(* Logix 5000 project; controller UOWHF_Vary Emulate 5570 rev 30.12; software revision 30.00; part 13 of 13 *)
(* tags used below, declared in another part *)
   UOWHF_Add_c : DINT;
   UOWHF_i : DINT;
   UOWHF_InputLen : DINT;
   UOWHF_InputMaxInd : DINT;
   UOWHF_Msg : DINT[16];
   UOWHF_OutputMaxInd : DINT;
   UOWHF_Result : DINT[17];
   UOWHF_Vary_BlkNum : DINT;
   UOWHF_Vary_i : DINT;
   UOWHF_Vary_j : DINT;
   UOWHF_Vary_Message : DINT[512];
   UOWHF_Vary_MsgLen : DINT;
   UOWHF_Vary_z : DINT;
   UOWHF_VaryLen : DINT;
   UOWHF_Ver : DINT;
(* MainProgram, continued *)

   		UOWHF_Add_c.7:=UOWHF_Result[7].31;
   		UOWHF_Result[7].31:=0;
   		UOWHF_Result[8]:=UOWHF_Result[8] + 1529564597+UOWHF_Add_c;
   		UOWHF_Add_c.8:=UOWHF_Result[8].31;
   		UOWHF_Result[8].31:=0;
   	End_If;
   	If UOWHF_Msg[15].[5] Then
   		UOWHF_Result[0]:=UOWHF_Result[0] + 534622081+UOWHF_Add_c;
   		UOWHF_Add_c.0:=UOWHF_Result[0].31;
   		UOWHF_Result[0].31:=0;
   		UOWHF_Result[1]:=UOWHF_Result[1] + 1054997605+UOWHF_Add_c;
   		UOWHF_Add_c.1:=UOWHF_Result[1].31;
   		UOWHF_Result[1].31:=0;
   		UOWHF_Result[2]:=UOWHF_Result[2] + 944898288+UOWHF_Add_c;
   		UOWHF_Add_c.2:=UOWHF_Result[2].31;
   		UOWHF_Result[2].31:=0;
   		UOWHF_Result[3]:=UOWHF_Result[3] + 811676453+UOWHF_Add_c;
   		UOWHF_Add_c.3:=UOWHF_Result[3].31;
   		UOWHF_Result[3].31:=0;
   		UOWHF_Result[4]:=UOWHF_Result[4] + 1761848356+UOWHF_Add_c;
   		UOWHF_Add_c.4:=UOWHF_Result[4].31;
   		UOWHF_Result[4].31:=0;
   		UOWHF_Result[5]:=UOWHF_Result[5] + 163403387+UOWHF_Add_c;
   		UOWHF_Add_c.5:=UOWHF_Result[5].31;
   		UOWHF_Result[5].31:=0;
   		UOWHF_Result[6]:=UOWHF_Result[6] + 606196183+UOWHF_Add_c;
   		UOWHF_Add_c.6:=UOWHF_Result[6].31;
   		UOWHF_Result[6].31:=0;
   		UOWHF_Result[7]:=UOWHF_Result[7] + 2030634477+UOWHF_Add_c;
   		UOWHF_Add_c.7:=UOWHF_Result[7].31;
   		UOWHF_Result[7].31:=0;
   		UOWHF_Result[8]:=UOWHF_Result[8] + 457492181+UOWHF_Add_c;
   		UOWHF_Add_c.8:=UOWHF_Result[8].31;
   		UOWHF_Result[8].31:=0;
   	End_If;
   	If UOWHF_Msg[15].[6] Then
   		UOWHF_Result[0]:=UOWHF_Result[0] + 1563595876+UOWHF_Add_c;
   		UOWHF_Add_c.0:=UOWHF_Result[0].31;
   		UOWHF_Result[0].31:=0;
   		UOWHF_Result[1]:=UOWHF_Result[1] + 921060794+UOWHF_Add_c;
   		UOWHF_Add_c.1:=UOWHF_Result[1].31;
   		UOWHF_Result[1].31:=0;
   		UOWHF_Result[2]:=UOWHF_Result[2] + 1052970481+UOWHF_Add_c;
   		UOWHF_Add_c.2:=UOWHF_Result[2].31;
   		UOWHF_Result[2].31:=0;
   		UOWHF_Result[3]:=UOWHF_Result[3] + 657088809+UOWHF_Add_c;
   		UOWHF_Add_c.3:=UOWHF_Result[3].31;
   		UOWHF_Result[3].31:=0;
   		UOWHF_Result[4]:=UOWHF_Result[4] + 107170927+UOWHF_Add_c;
   		UOWHF_Add_c.4:=UOWHF_Result[4].31;
   		UOWHF_Result[4].31:=0;
   		UOWHF_Result[5]:=UOWHF_Result[5] + 1430973014+UOWHF_Add_c;
   		UOWHF_Add_c.5:=UOWHF_Result[5].31;
   		UOWHF_Result[5].31:=0;
   		UOWHF_Result[6]:=UOWHF_Result[6] + 454401316+UOWHF_Add_c;
   		UOWHF_Add_c.6:=UOWHF_Result[6].31;
   		UOWHF_Result[6].31:=0;
   		UOWHF_Result[7]:=UOWHF_Result[7] + 395129130+UOWHF_Add_c;
   		UOWHF_Add_c.7:=UOWHF_Result[7].31;
   		UOWHF_Result[7].31:=0;
   		UOWHF_Result[8]:=UOWHF_Result[8] + 1072078032+UOWHF_Add_c;
   		UOWHF_Add_c.8:=UOWHF_Result[8].31;
   		UOWHF_Result[8].31:=0;
   	End_If;
   	If UOWHF_Msg[15].[7] Then
   		UOWHF_Result[0]:=UOWHF_Result[0] + 1403391658+UOWHF_Add_c;
   		UOWHF_Add_c.0:=UOWHF_Result[0].31;
   		UOWHF_Result[0].31:=0;
   		UOWHF_Result[1]:=UOWHF_Result[1] + 1796223182+UOWHF_Add_c;
   		UOWHF_Add_c.1:=UOWHF_Result[1].31;
   		UOWHF_Result[1].31:=0;
   		UOWHF_Result[2]:=UOWHF_Result[2] + 960792761+UOWHF_Add_c;
   		UOWHF_Add_c.2:=UOWHF_Result[2].31;
   		UOWHF_Result[2].31:=0;
   		UOWHF_Result[3]:=UOWHF_Result[3] + 288040454+UOWHF_Add_c;
   		UOWHF_Add_c.3:=UOWHF_Result[3].31;
   		UOWHF_Result[3].31:=0;
   		UOWHF_Result[4]:=UOWHF_Result[4] + 356603480+UOWHF_Add_c;
   		UOWHF_Add_c.4:=UOWHF_Result[4].31;
   		UOWHF_Result[4].31:=0;
   		UOWHF_Result[5]:=UOWHF_Result[5] + 1694776766+UOWHF_Add_c;
   		UOWHF_Add_c.5:=UOWHF_Result[5].31;
   		UOWHF_Result[5].31:=0;
   		UOWHF_Result[6]:=UOWHF_Result[6] + 1001613380+UOWHF_Add_c;
   		UOWHF_Add_c.6:=UOWHF_Result[6].31;
   		UOWHF_Result[6].31:=0;
   		UOWHF_Result[7]:=UOWHF_Result[7] + 1296327921+UOWHF_Add_c;
   		UOWHF_Add_c.7:=UOWHF_Result[7].31;
   		UOWHF_Result[7].31:=0;
   		UOWHF_Result[8]:=UOWHF_Result[8] + 1853983857+UOWHF_Add_c;
   		UOWHF_Add_c.8:=UOWHF_Result[8].31;
   		UOWHF_Result[8].31:=0;
   	End_If;
   	If UOWHF_Msg[15].[8] Then
   		UOWHF_Result[0]:=UOWHF_Result[0] + 1265129415+UOWHF_Add_c;
   		UOWHF_Add_c.0:=UOWHF_Result[0].31;
   		UOWHF_Result[0].31:=0;
   		UOWHF_Result[1]:=UOWHF_Result[1] + 568656446+UOWHF_Add_c;
   		UOWHF_Add_c.1:=UOWHF_Result[1].31;
   		UOWHF_Result[1].31:=0;
   		UOWHF_Result[2]:=UOWHF_Result[2] + 1035914428+UOWHF_Add_c;
   		UOWHF_Add_c.2:=UOWHF_Result[2].31;
   		UOWHF_Result[2].31:=0;
   		UOWHF_Result[3]:=UOWHF_Result[3] + 1838467801+UOWHF_Add_c;
   		UOWHF_Add_c.3:=UOWHF_Result[3].31;
   		UOWHF_Result[3].31:=0;
   		UOWHF_Result[4]:=UOWHF_Result[4] + 852571844+UOWHF_Add_c;
   		UOWHF_Add_c.4:=UOWHF_Result[4].31;
   		UOWHF_Result[4].31:=0;
   		UOWHF_Result[5]:=UOWHF_Result[5] + 811437709+UOWHF_Add_c;
   		UOWHF_Add_c.5:=UOWHF_Result[5].31;
   		UOWHF_Result[5].31:=0;
   		UOWHF_Result[6]:=UOWHF_Result[6] + 2110578431+UOWHF_Add_c;
   		UOWHF_Add_c.6:=UOWHF_Result[6].31;
   		UOWHF_Result[6].31:=0;
   		UOWHF_Result[7]:=UOWHF_Result[7] + 1083369967+UOWHF_Add_c;
   		UOWHF_Add_c.7:=UOWHF_Result[7].31;
   		UOWHF_Result[7].31:=0;
   		UOWHF_Result[8]:=UOWHF_Result[8] + 1040887567+UOWHF_Add_c;
   		UOWHF_Add_c.8:=UOWHF_Result[8].31;
   		UOWHF_Result[8].31:=0;
   	End_If;
   	If UOWHF_Msg[15].[9] Then
   		UOWHF_Result[0]:=UOWHF_Result[0] + 1883016459+UOWHF_Add_c;
   		UOWHF_Add_c.0:=UOWHF_Result[0].31;
   		UOWHF_Result[0].31:=0;
   		UOWHF_Result[1]:=UOWHF_Result[1] + 1109215782+UOWHF_Add_c;
   		UOWHF_Add_c.1:=UOWHF_Result[1].31;
   		UOWHF_Result[1].31:=0;
   		UOWHF_Result[2]:=UOWHF_Result[2] + 692572348+UOWHF_Add_c;
   		UOWHF_Add_c.2:=UOWHF_Result[2].31;
   		UOWHF_Result[2].31:=0;
   		UOWHF_Result[3]:=UOWHF_Result[3] + 357248589+UOWHF_Add_c;
   		UOWHF_Add_c.3:=UOWHF_Result[3].31;
   		UOWHF_Result[3].31:=0;
   		UOWHF_Result[4]:=UOWHF_Result[4] + 495139913+UOWHF_Add_c;
   		UOWHF_Add_c.4:=UOWHF_Result[4].31;
   		UOWHF_Result[4].31:=0;
   		UOWHF_Result[5]:=UOWHF_Result[5] + 1972425862+UOWHF_Add_c;
   		UOWHF_Add_c.5:=UOWHF_Result[5].31;
   		UOWHF_Result[5].31:=0;
   		UOWHF_Result[6]:=UOWHF_Result[6] + 1336574867+UOWHF_Add_c;
   		UOWHF_Add_c.6:=UOWHF_Result[6].31;
   		UOWHF_Result[6].31:=0;
   		UOWHF_Result[7]:=UOWHF_Result[7] + 286906005+UOWHF_Add_c;
   		UOWHF_Add_c.7:=UOWHF_Result[7].31;
   		UOWHF_Result[7].31:=0;
   		UOWHF_Result[8]:=UOWHF_Result[8] + 935997948+UOWHF_Add_c;
   		UOWHF_Add_c.8:=UOWHF_Result[8].31;
   		UOWHF_Result[8].31:=0;
   	End_If;
   	If UOWHF_Msg[15].[10] Then
   		UOWHF_Result[0]:=UOWHF_Result[0] + 406811790+UOWHF_Add_c;
   		UOWHF_Add_c.0:=UOWHF_Result[0].31;
   		UOWHF_Result[0].31:=0;
   		UOWHF_Result[1]:=UOWHF_Result[1] + 1667294919+UOWHF_Add_c;
   		UOWHF_Add_c.1:=UOWHF_Result[1].31;
   		UOWHF_Result[1].31:=0;
   		UOWHF_Result[2]:=UOWHF_Result[2] + 2033524595+UOWHF_Add_c;
   		UOWHF_Add_c.2:=UOWHF_Result[2].31;
   		UOWHF_Result[2].31:=0;
   		UOWHF_Result[3]:=UOWHF_Result[3] + 1349255026+UOWHF_Add_c;
   		UOWHF_Add_c.3:=UOWHF_Result[3].31;
   		UOWHF_Result[3].31:=0;
   		UOWHF_Result[4]:=UOWHF_Result[4] + 10415662+UOWHF_Add_c;
   		UOWHF_Add_c.4:=UOWHF_Result[4].31;
   		UOWHF_Result[4].31:=0;
   		UOWHF_Result[5]:=UOWHF_Result[5] + 2068656448+UOWHF_Add_c;
   		UOWHF_Add_c.5:=UOWHF_Result[5].31;
   		UOWHF_Result[5].31:=0;
   		UOWHF_Result[6]:=UOWHF_Result[6] + 719617830+UOWHF_Add_c;
   		UOWHF_Add_c.6:=UOWHF_Result[6].31;
   		UOWHF_Result[6].31:=0;
   		UOWHF_Result[7]:=UOWHF_Result[7] + 867653174+UOWHF_Add_c;
   		UOWHF_Add_c.7:=UOWHF_Result[7].31;
   		UOWHF_Result[7].31:=0;
   		UOWHF_Result[8]:=UOWHF_Result[8] + 1934472738+UOWHF_Add_c;
   		UOWHF_Add_c.8:=UOWHF_Result[8].31;
   		UOWHF_Result[8].31:=0;
   	End_If;
   	If UOWHF_Msg[15].[11] Then
   		UOWHF_Result[0]:=UOWHF_Result[0] + 165633326+UOWHF_Add_c;
   		UOWHF_Add_c.0:=UOWHF_Result[0].31;
   		UOWHF_Result[0].31:=0;
   		UOWHF_Result[1]:=UOWHF_Result[1] + 53652767+UOWHF_Add_c;
   		UOWHF_Add_c.1:=UOWHF_Result[1].31;
   		UOWHF_Result[1].31:=0;
   		UOWHF_Result[2]:=UOWHF_Result[2] + 1574797324+UOWHF_Add_c;
   		UOWHF_Add_c.2:=UOWHF_Result[2].31;
   		UOWHF_Result[2].31:=0;
   		UOWHF_Result[3]:=UOWHF_Result[3] + 1336775684+UOWHF_Add_c;
   		UOWHF_Add_c.3:=UOWHF_Result[3].31;
   		UOWHF_Result[3].31:=0;
   		UOWHF_Result[4]:=UOWHF_Result[4] + 1894121389+UOWHF_Add_c;
   		UOWHF_Add_c.4:=UOWHF_Result[4].31;
   		UOWHF_Result[4].31:=0;
   		UOWHF_Result[5]:=UOWHF_Result[5] + 1658923569+UOWHF_Add_c;
   		UOWHF_Add_c.5:=UOWHF_Result[5].31;
   		UOWHF_Result[5].31:=0;
   		UOWHF_Result[6]:=UOWHF_Result[6] + 1195345328+UOWHF_Add_c;
   		UOWHF_Add_c.6:=UOWHF_Result[6].31;
   		UOWHF_Result[6].31:=0;
   		UOWHF_Result[7]:=UOWHF_Result[7] + 1912811518+UOWHF_Add_c;
   		UOWHF_Add_c.7:=UOWHF_Result[7].31;
   		UOWHF_Result[7].31:=0;
   		UOWHF_Result[8]:=UOWHF_Result[8] + 826695963+UOWHF_Add_c;
   		UOWHF_Add_c.8:=UOWHF_Result[8].31;
   		UOWHF_Result[8].31:=0;
   	End_If;
   	If UOWHF_Msg[15].[12] Then
   		UOWHF_Result[0]:=UOWHF_Result[0] + 1033530810+UOWHF_Add_c;
   		UOWHF_Add_c.0:=UOWHF_Result[0].31;
   		UOWHF_Result[0].31:=0;
   		UOWHF_Result[1]:=UOWHF_Result[1] + 449682606+UOWHF_Add_c;
   		UOWHF_Add_c.1:=UOWHF_Result[1].31;
   		UOWHF_Result[1].31:=0;
   		UOWHF_Result[2]:=UOWHF_Result[2] + 1100837890+UOWHF_Add_c;
   		UOWHF_Add_c.2:=UOWHF_Result[2].31;
   		UOWHF_Result[2].31:=0;
   		UOWHF_Result[3]:=UOWHF_Result[3] + 721973923+UOWHF_Add_c;
   		UOWHF_Add_c.3:=UOWHF_Result[3].31;
   		UOWHF_Result[3].31:=0;
   		UOWHF_Result[4]:=UOWHF_Result[4] + 2071465357+UOWHF_Add_c;
   		UOWHF_Add_c.4:=UOWHF_Result[4].31;
   		UOWHF_Result[4].31:=0;
   		UOWHF_Result[5]:=UOWHF_Result[5] + 514392075+UOWHF_Add_c;
   		UOWHF_Add_c.5:=UOWHF_Result[5].31;
   		UOWHF_Result[5].31:=0;
   		UOWHF_Result[6]:=UOWHF_Result[6] + 241897951+UOWHF_Add_c;
   		UOWHF_Add_c.6:=UOWHF_Result[6].31;
   		UOWHF_Result[6].31:=0;
   		UOWHF_Result[7]:=UOWHF_Result[7] + 1971083301+UOWHF_Add_c;
   		UOWHF_Add_c.7:=UOWHF_Result[7].31;
   		UOWHF_Result[7].31:=0;
   		UOWHF_Result[8]:=UOWHF_Result[8] + 326292913+UOWHF_Add_c;
   		UOWHF_Add_c.8:=UOWHF_Result[8].31;
   		UOWHF_Result[8].31:=0;
   	End_If;
   	If UOWHF_Msg[15].[13] Then
   		UOWHF_Result[0]:=UOWHF_Result[0] + 827872352+UOWHF_Add_c;
   		UOWHF_Add_c.0:=UOWHF_Result[0].31;
   		UOWHF_Result[0].31:=0;
   		UOWHF_Result[1]:=UOWHF_Result[1] + 1501229297+UOWHF_Add_c;
   		UOWHF_Add_c.1:=UOWHF_Result[1].31;
   		UOWHF_Result[1].31:=0;
   		UOWHF_Result[2]:=UOWHF_Result[2] + 140749544+UOWHF_Add_c;
   		UOWHF_Add_c.2:=UOWHF_Result[2].31;
   		UOWHF_Result[2].31:=0;
   		UOWHF_Result[3]:=UOWHF_Result[3] + 604970260+UOWHF_Add_c;
   		UOWHF_Add_c.3:=UOWHF_Result[3].31;
   		UOWHF_Result[3].31:=0;
   		UOWHF_Result[4]:=UOWHF_Result[4] + 1399783902+UOWHF_Add_c;
   		UOWHF_Add_c.4:=UOWHF_Result[4].31;
   		UOWHF_Result[4].31:=0;
   		UOWHF_Result[5]:=UOWHF_Result[5] + 697715354+UOWHF_Add_c;
   		UOWHF_Add_c.5:=UOWHF_Result[5].31;
   		UOWHF_Result[5].31:=0;
   		UOWHF_Result[6]:=UOWHF_Result[6] + 1132588250+UOWHF_Add_c;
   		UOWHF_Add_c.6:=UOWHF_Result[6].31;
   		UOWHF_Result[6].31:=0;
   		UOWHF_Result[7]:=UOWHF_Result[7] + 1508151598+UOWHF_Add_c;
   		UOWHF_Add_c.7:=UOWHF_Result[7].31;
   		UOWHF_Result[7].31:=0;
   		UOWHF_Result[8]:=UOWHF_Result[8] + 575502560+UOWHF_Add_c;
   		UOWHF_Add_c.8:=UOWHF_Result[8].31;
   		UOWHF_Result[8].31:=0;
   	End_If;
   	If UOWHF_Msg[15].[14] Then
   		UOWHF_Result[0]:=UOWHF_Result[0] + 1928657576+UOWHF_Add_c;
   		UOWHF_Add_c.0:=UOWHF_Result[0].31;
   		UOWHF_Result[0].31:=0;
   		UOWHF_Result[1]:=UOWHF_Result[1] + 1105884606+UOWHF_Add_c;
   		UOWHF_Add_c.1:=UOWHF_Result[1].31;
   		UOWHF_Result[1].31:=0;
   		UOWHF_Result[2]:=UOWHF_Result[2] + 106499913+UOWHF_Add_c;
   		UOWHF_Add_c.2:=UOWHF_Result[2].31;
   		UOWHF_Result[2].31:=0;
   		UOWHF_Result[3]:=UOWHF_Result[3] + 1490777468+UOWHF_Add_c;
   		UOWHF_Add_c.3:=UOWHF_Result[3].31;
   		UOWHF_Result[3].31:=0;
   		UOWHF_Result[4]:=UOWHF_Result[4] + 76282737+UOWHF_Add_c;
   		UOWHF_Add_c.4:=UOWHF_Result[4].31;
   		UOWHF_Result[4].31:=0;
   		UOWHF_Result[5]:=UOWHF_Result[5] + 524228130+UOWHF_Add_c;
   		UOWHF_Add_c.5:=UOWHF_Result[5].31;
   		UOWHF_Result[5].31:=0;
   		UOWHF_Result[6]:=UOWHF_Result[6] + 1228552707+UOWHF_Add_c;
   		UOWHF_Add_c.6:=UOWHF_Result[6].31;
   		UOWHF_Result[6].31:=0;
   		UOWHF_Result[7]:=UOWHF_Result[7] + 1666564749+UOWHF_Add_c;
   		UOWHF_Add_c.7:=UOWHF_Result[7].31;
   		UOWHF_Result[7].31:=0;
   		UOWHF_Result[8]:=UOWHF_Result[8] + 268528645+UOWHF_Add_c;
   		UOWHF_Add_c.8:=UOWHF_Result[8].31;
   		UOWHF_Result[8].31:=0;
   	End_If;
   	If UOWHF_Msg[15].[15] Then
   		UOWHF_Result[0]:=UOWHF_Result[0] + 1961791867+UOWHF_Add_c;
   		UOWHF_Add_c.0:=UOWHF_Result[0].31;
   		UOWHF_Result[0].31:=0;
   		UOWHF_Result[1]:=UOWHF_Result[1] + 952816348+UOWHF_Add_c;
   		UOWHF_Add_c.1:=UOWHF_Result[1].31;
   		UOWHF_Result[1].31:=0;
   		UOWHF_Result[2]:=UOWHF_Result[2] + 136661959+UOWHF_Add_c;
   		UOWHF_Add_c.2:=UOWHF_Result[2].31;
   		UOWHF_Result[2].31:=0;
   		UOWHF_Result[3]:=UOWHF_Result[3] + 178536398+UOWHF_Add_c;
   		UOWHF_Add_c.3:=UOWHF_Result[3].31;
   		UOWHF_Result[3].31:=0;
   		UOWHF_Result[4]:=UOWHF_Result[4] + 1561223972+UOWHF_Add_c;
   		UOWHF_Add_c.4:=UOWHF_Result[4].31;
   		UOWHF_Result[4].31:=0;
   		UOWHF_Result[5]:=UOWHF_Result[5] + 1593802136+UOWHF_Add_c;
   		UOWHF_Add_c.5:=UOWHF_Result[5].31;
   		UOWHF_Result[5].31:=0;
   		UOWHF_Result[6]:=UOWHF_Result[6] + 1412200351+UOWHF_Add_c;
   		UOWHF_Add_c.6:=UOWHF_Result[6].31;
   		UOWHF_Result[6].31:=0;
   		UOWHF_Result[7]:=UOWHF_Result[7] + 1568670030+UOWHF_Add_c;
   		UOWHF_Add_c.7:=UOWHF_Result[7].31;
   		UOWHF_Result[7].31:=0;
   		UOWHF_Result[8]:=UOWHF_Result[8] + 967013106+UOWHF_Add_c;
   		UOWHF_Add_c.8:=UOWHF_Result[8].31;
   		UOWHF_Result[8].31:=0;
   	End_If;
   	If UOWHF_Msg[15].[16] Then
   		UOWHF_Result[0]:=UOWHF_Result[0] + 169683100+UOWHF_Add_c;
   		UOWHF_Add_c.0:=UOWHF_Result[0].31;
   		UOWHF_Result[0].31:=0;
   		UOWHF_Result[1]:=UOWHF_Result[1] + 570495153+UOWHF_Add_c;
   		UOWHF_Add_c.1:=UOWHF_Result[1].31;
   		UOWHF_Result[1].31:=0;
   		UOWHF_Result[2]:=UOWHF_Result[2] + 1798228575+UOWHF_Add_c;
   		UOWHF_Add_c.2:=UOWHF_Result[2].31;
   		UOWHF_Result[2].31:=0;
   		UOWHF_Result[3]:=UOWHF_Result[3] + 1246241515+UOWHF_Add_c;
   		UOWHF_Add_c.3:=UOWHF_Result[3].31;
   		UOWHF_Result[3].31:=0;
   		UOWHF_Result[4]:=UOWHF_Result[4] + 2135845928+UOWHF_Add_c;
   		UOWHF_Add_c.4:=UOWHF_Result[4].31;
   		UOWHF_Result[4].31:=0;
   		UOWHF_Result[5]:=UOWHF_Result[5] + 456024302+UOWHF_Add_c;
   		UOWHF_Add_c.5:=UOWHF_Result[5].31;
   		UOWHF_Result[5].31:=0;
   		UOWHF_Result[6]:=UOWHF_Result[6] + 1289737613+UOWHF_Add_c;
   		UOWHF_Add_c.6:=UOWHF_Result[6].31;
   		UOWHF_Result[6].31:=0;
   		UOWHF_Result[7]:=UOWHF_Result[7] + 1705301408+UOWHF_Add_c;
   		UOWHF_Add_c.7:=UOWHF_Result[7].31;
   		UOWHF_Result[7].31:=0;
   		UOWHF_Result[8]:=UOWHF_Result[8] + 1734663976+UOWHF_Add_c;
   		UOWHF_Add_c.8:=UOWHF_Result[8].31;
   		UOWHF_Result[8].31:=0;
   	End_If;
   	If UOWHF_Msg[15].[17] Then
   		UOWHF_Result[0]:=UOWHF_Result[0] + 983372193+UOWHF_Add_c;
   		UOWHF_Add_c.0:=UOWHF_Result[0].31;
   		UOWHF_Result[0].31:=0;
   		UOWHF_Result[1]:=UOWHF_Result[1] + 638884961+UOWHF_Add_c;
   		UOWHF_Add_c.1:=UOWHF_Result[1].31;
   		UOWHF_Result[1].31:=0;
   		UOWHF_Result[2]:=UOWHF_Result[2] + 1694858606+UOWHF_Add_c;
   		UOWHF_Add_c.2:=UOWHF_Result[2].31;
   		UOWHF_Result[2].31:=0;
   		UOWHF_Result[3]:=UOWHF_Result[3] + 284670684+UOWHF_Add_c;
   		UOWHF_Add_c.3:=UOWHF_Result[3].31;
   		UOWHF_Result[3].31:=0;
   		UOWHF_Result[4]:=UOWHF_Result[4] + 25547865+UOWHF_Add_c;
   		UOWHF_Add_c.4:=UOWHF_Result[4].31;
   		UOWHF_Result[4].31:=0;
   		UOWHF_Result[5]:=UOWHF_Result[5] + 1037524440+UOWHF_Add_c;
   		UOWHF_Add_c.5:=UOWHF_Result[5].31;
   		UOWHF_Result[5].31:=0;
   		UOWHF_Result[6]:=UOWHF_Result[6] + 1634584801+UOWHF_Add_c;
   		UOWHF_Add_c.6:=UOWHF_Result[6].31;
   		UOWHF_Result[6].31:=0;
   		UOWHF_Result[7]:=UOWHF_Result[7] + 818446873+UOWHF_Add_c;
   		UOWHF_Add_c.7:=UOWHF_Result[7].31;
   		UOWHF_Result[7].31:=0;
   		UOWHF_Result[8]:=UOWHF_Result[8] + 1700629153+UOWHF_Add_c;
   		UOWHF_Add_c.8:=UOWHF_Result[8].31;
   		UOWHF_Result[8].31:=0;
   	End_If;
   	If UOWHF_Msg[15].[18] Then
   		UOWHF_Result[0]:=UOWHF_Result[0] + 78321704+UOWHF_Add_c;
   		UOWHF_Add_c.0:=UOWHF_Result[0].31;
   		UOWHF_Result[0].31:=0;
   		UOWHF_Result[1]:=UOWHF_Result[1] + 1937348808+UOWHF_Add_c;
   		UOWHF_Add_c.1:=UOWHF_Result[1].31;
   		UOWHF_Result[1].31:=0;
   		UOWHF_Result[2]:=UOWHF_Result[2] + 130465258+UOWHF_Add_c;
   		UOWHF_Add_c.2:=UOWHF_Result[2].31;
   		UOWHF_Result[2].31:=0;
   		UOWHF_Result[3]:=UOWHF_Result[3] + 1461020702+UOWHF_Add_c;
   		UOWHF_Add_c.3:=UOWHF_Result[3].31;
   		UOWHF_Result[3].31:=0;
   		UOWHF_Result[4]:=UOWHF_Result[4] + 1957110397+UOWHF_Add_c;
   		UOWHF_Add_c.4:=UOWHF_Result[4].31;
   		UOWHF_Result[4].31:=0;
   		UOWHF_Result[5]:=UOWHF_Result[5] + 1790059909+UOWHF_Add_c;
   		UOWHF_Add_c.5:=UOWHF_Result[5].31;
   		UOWHF_Result[5].31:=0;
   		UOWHF_Result[6]:=UOWHF_Result[6] + 857304694+UOWHF_Add_c;
   		UOWHF_Add_c.6:=UOWHF_Result[6].31;
   		UOWHF_Result[6].31:=0;
   		UOWHF_Result[7]:=UOWHF_Result[7] + 1509154065+UOWHF_Add_c;
   		UOWHF_Add_c.7:=UOWHF_Result[7].31;
   		UOWHF_Result[7].31:=0;
   		UOWHF_Result[8]:=UOWHF_Result[8] + 1157248973+UOWHF_Add_c;
   		UOWHF_Add_c.8:=UOWHF_Result[8].31;
   		UOWHF_Result[8].31:=0;
   	End_If;
   	If UOWHF_Msg[15].[19] Then
   		UOWHF_Result[0]:=UOWHF_Result[0] + 552710964+UOWHF_Add_c;
   		UOWHF_Add_c.0:=UOWHF_Result[0].31;
   		UOWHF_Result[0].31:=0;
   		UOWHF_Result[1]:=UOWHF_Result[1] + 1128382434+UOWHF_Add_c;
   		UOWHF_Add_c.1:=UOWHF_Result[1].31;
   		UOWHF_Result[1].31:=0;
   		UOWHF_Result[2]:=UOWHF_Result[2] + 1867237623+UOWHF_Add_c;
   		UOWHF_Add_c.2:=UOWHF_Result[2].31;
   		UOWHF_Result[2].31:=0;
   		UOWHF_Result[3]:=UOWHF_Result[3] + 2146368693+UOWHF_Add_c;
   		UOWHF_Add_c.3:=UOWHF_Result[3].31;
   		UOWHF_Result[3].31:=0;
   		UOWHF_Result[4]:=UOWHF_Result[4] + 1142566885+UOWHF_Add_c;
   		UOWHF_Add_c.4:=UOWHF_Result[4].31;
   		UOWHF_Result[4].31:=0;
   		UOWHF_Result[5]:=UOWHF_Result[5] + 861229388+UOWHF_Add_c;
   		UOWHF_Add_c.5:=UOWHF_Result[5].31;
   		UOWHF_Result[5].31:=0;
   		UOWHF_Result[6]:=UOWHF_Result[6] + 698199324+UOWHF_Add_c;
   		UOWHF_Add_c.6:=UOWHF_Result[6].31;
   		UOWHF_Result[6].31:=0;
   		UOWHF_Result[7]:=UOWHF_Result[7] + 2095517647+UOWHF_Add_c;
   		UOWHF_Add_c.7:=UOWHF_Result[7].31;
   		UOWHF_Result[7].31:=0;
   		UOWHF_Result[8]:=UOWHF_Result[8] + 1174160295+UOWHF_Add_c;
   		UOWHF_Add_c.8:=UOWHF_Result[8].31;
   		UOWHF_Result[8].31:=0;
   	End_If;
   	If UOWHF_Msg[15].[20] Then
   		UOWHF_Result[0]:=UOWHF_Result[0] + 1585620937+UOWHF_Add_c;
   		UOWHF_Add_c.0:=UOWHF_Result[0].31;
   		UOWHF_Result[0].31:=0;
   		UOWHF_Result[1]:=UOWHF_Result[1] + 325026118+UOWHF_Add_c;
   		UOWHF_Add_c.1:=UOWHF_Result[1].31;
   		UOWHF_Result[1].31:=0;
   		UOWHF_Result[2]:=UOWHF_Result[2] + 738436433+UOWHF_Add_c;
   		UOWHF_Add_c.2:=UOWHF_Result[2].31;
   		UOWHF_Result[2].31:=0;
   		UOWHF_Result[3]:=UOWHF_Result[3] + 1422046785+UOWHF_Add_c;
   		UOWHF_Add_c.3:=UOWHF_Result[3].31;
   		UOWHF_Result[3].31:=0;
   		UOWHF_Result[4]:=UOWHF_Result[4] + 1969896335+UOWHF_Add_c;
   		UOWHF_Add_c.4:=UOWHF_Result[4].31;
   		UOWHF_Result[4].31:=0;
   		UOWHF_Result[5]:=UOWHF_Result[5] + 191628607+UOWHF_Add_c;
   		UOWHF_Add_c.5:=UOWHF_Result[5].31;
   		UOWHF_Result[5].31:=0;
   		UOWHF_Result[6]:=UOWHF_Result[6] + 1650724515+UOWHF_Add_c;
   		UOWHF_Add_c.6:=UOWHF_Result[6].31;
   		UOWHF_Result[6].31:=0;
   		UOWHF_Result[7]:=UOWHF_Result[7] + 361882123+UOWHF_Add_c;
   		UOWHF_Add_c.7:=UOWHF_Result[7].31;
   		UOWHF_Result[7].31:=0;
   		UOWHF_Result[8]:=UOWHF_Result[8] + 989278147+UOWHF_Add_c;
   		UOWHF_Add_c.8:=UOWHF_Result[8].31;
   		UOWHF_Result[8].31:=0;
   	End_If;
   	If UOWHF_Msg[15].[21] Then
   		UOWHF_Result[0]:=UOWHF_Result[0] + 1462556247+UOWHF_Add_c;
   		UOWHF_Add_c.0:=UOWHF_Result[0].31;
   		UOWHF_Result[0].31:=0;
   		UOWHF_Result[1]:=UOWHF_Result[1] + 99576052+UOWHF_Add_c;
   		UOWHF_Add_c.1:=UOWHF_Result[1].31;
   		UOWHF_Result[1].31:=0;
   		UOWHF_Result[2]:=UOWHF_Result[2] + 202621392+UOWHF_Add_c;
   		UOWHF_Add_c.2:=UOWHF_Result[2].31;
   		UOWHF_Result[2].31:=0;
   		UOWHF_Result[3]:=UOWHF_Result[3] + 67765093+UOWHF_Add_c;
   		UOWHF_Add_c.3:=UOWHF_Result[3].31;
   		UOWHF_Result[3].31:=0;
   		UOWHF_Result[4]:=UOWHF_Result[4] + 1059801784+UOWHF_Add_c;
   		UOWHF_Add_c.4:=UOWHF_Result[4].31;
   		UOWHF_Result[4].31:=0;
   		UOWHF_Result[5]:=UOWHF_Result[5] + 1364564603+UOWHF_Add_c;
   		UOWHF_Add_c.5:=UOWHF_Result[5].31;
   		UOWHF_Result[5].31:=0;
   		UOWHF_Result[6]:=UOWHF_Result[6] + 1133940393+UOWHF_Add_c;
   		UOWHF_Add_c.6:=UOWHF_Result[6].31;
   		UOWHF_Result[6].31:=0;
   		UOWHF_Result[7]:=UOWHF_Result[7] + 740275323+UOWHF_Add_c;
   		UOWHF_Add_c.7:=UOWHF_Result[7].31;
   		UOWHF_Result[7].31:=0;
   		UOWHF_Result[8]:=UOWHF_Result[8] + 211656668+UOWHF_Add_c;
   		UOWHF_Add_c.8:=UOWHF_Result[8].31;
   		UOWHF_Result[8].31:=0;
   	End_If;
   	If UOWHF_Msg[15].[22] Then
   		UOWHF_Result[0]:=UOWHF_Result[0] + 940319263+UOWHF_Add_c;
   		UOWHF_Add_c.0:=UOWHF_Result[0].31;
   		UOWHF_Result[0].31:=0;
   		UOWHF_Result[1]:=UOWHF_Result[1] + 1171691104+UOWHF_Add_c;
   		UOWHF_Add_c.1:=UOWHF_Result[1].31;
   		UOWHF_Result[1].31:=0;
   		UOWHF_Result[2]:=UOWHF_Result[2] + 1620828792+UOWHF_Add_c;
   		UOWHF_Add_c.2:=UOWHF_Result[2].31;
   		UOWHF_Result[2].31:=0;
   		UOWHF_Result[3]:=UOWHF_Result[3] + 889659934+UOWHF_Add_c;
   		UOWHF_Add_c.3:=UOWHF_Result[3].31;
   		UOWHF_Result[3].31:=0;
   		UOWHF_Result[4]:=UOWHF_Result[4] + 246769229+UOWHF_Add_c;
   		UOWHF_Add_c.4:=UOWHF_Result[4].31;
   		UOWHF_Result[4].31:=0;
   		UOWHF_Result[5]:=UOWHF_Result[5] + 1871507547+UOWHF_Add_c;
   		UOWHF_Add_c.5:=UOWHF_Result[5].31;
   		UOWHF_Result[5].31:=0;
   		UOWHF_Result[6]:=UOWHF_Result[6] + 1111223933+UOWHF_Add_c;
   		UOWHF_Add_c.6:=UOWHF_Result[6].31;
   		UOWHF_Result[6].31:=0;
   		UOWHF_Result[7]:=UOWHF_Result[7] + 1590368283+UOWHF_Add_c;
   		UOWHF_Add_c.7:=UOWHF_Result[7].31;
   		UOWHF_Result[7].31:=0;
   		UOWHF_Result[8]:=UOWHF_Result[8] + 475158687+UOWHF_Add_c;
   		UOWHF_Add_c.8:=UOWHF_Result[8].31;
   		UOWHF_Result[8].31:=0;
   	End_If;
   	If UOWHF_Msg[15].[23] Then
   		UOWHF_Result[0]:=UOWHF_Result[0] + 1294958433+UOWHF_Add_c;
   		UOWHF_Add_c.0:=UOWHF_Result[0].31;
   		UOWHF_Result[0].31:=0;
   		UOWHF_Result[1]:=UOWHF_Result[1] + 815634209+UOWHF_Add_c;
   		UOWHF_Add_c.1:=UOWHF_Result[1].31;
   		UOWHF_Result[1].31:=0;
   		UOWHF_Result[2]:=UOWHF_Result[2] + 1757336081+UOWHF_Add_c;
   		UOWHF_Add_c.2:=UOWHF_Result[2].31;
   		UOWHF_Result[2].31:=0;
   		UOWHF_Result[3]:=UOWHF_Result[3] + 657179249+UOWHF_Add_c;
   		UOWHF_Add_c.3:=UOWHF_Result[3].31;
   		UOWHF_Result[3].31:=0;
   		UOWHF_Result[4]:=UOWHF_Result[4] + 1827267451+UOWHF_Add_c;
   		UOWHF_Add_c.4:=UOWHF_Result[4].31;
   		UOWHF_Result[4].31:=0;
   		UOWHF_Result[5]:=UOWHF_Result[5] + 374874832+UOWHF_Add_c;
   		UOWHF_Add_c.5:=UOWHF_Result[5].31;
   		UOWHF_Result[5].31:=0;
   		UOWHF_Result[6]:=UOWHF_Result[6] + 312266219+UOWHF_Add_c;
   		UOWHF_Add_c.6:=UOWHF_Result[6].31;
   		UOWHF_Result[6].31:=0;
   		UOWHF_Result[7]:=UOWHF_Result[7] + 1133795400+UOWHF_Add_c;
   		UOWHF_Add_c.7:=UOWHF_Result[7].31;
   		UOWHF_Result[7].31:=0;
   		UOWHF_Result[8]:=UOWHF_Result[8] + 932878339+UOWHF_Add_c;
   		UOWHF_Add_c.8:=UOWHF_Result[8].31;
   		UOWHF_Result[8].31:=0;
   	End_If;
   	If UOWHF_Msg[15].[24] Then
   		UOWHF_Result[0]:=UOWHF_Result[0] + 332648701+UOWHF_Add_c;
   		UOWHF_Add_c.0:=UOWHF_Result[0].31;
   		UOWHF_Result[0].31:=0;
   		UOWHF_Result[1]:=UOWHF_Result[1] + 85758604+UOWHF_Add_c;
   		UOWHF_Add_c.1:=UOWHF_Result[1].31;
   		UOWHF_Result[1].31:=0;
   		UOWHF_Result[2]:=UOWHF_Result[2] + 971705346+UOWHF_Add_c;
   		UOWHF_Add_c.2:=UOWHF_Result[2].31;
   		UOWHF_Result[2].31:=0;
   		UOWHF_Result[3]:=UOWHF_Result[3] + 1047049167+UOWHF_Add_c;
   		UOWHF_Add_c.3:=UOWHF_Result[3].31;
   		UOWHF_Result[3].31:=0;
   		UOWHF_Result[4]:=UOWHF_Result[4] + 1221582178+UOWHF_Add_c;
   		UOWHF_Add_c.4:=UOWHF_Result[4].31;
   		UOWHF_Result[4].31:=0;
   		UOWHF_Result[5]:=UOWHF_Result[5] + 1982046425+UOWHF_Add_c;
   		UOWHF_Add_c.5:=UOWHF_Result[5].31;
   		UOWHF_Result[5].31:=0;
   		UOWHF_Result[6]:=UOWHF_Result[6] + 2109992137+UOWHF_Add_c;
   		UOWHF_Add_c.6:=UOWHF_Result[6].31;
   		UOWHF_Result[6].31:=0;
   		UOWHF_Result[7]:=UOWHF_Result[7] + 1514276956+UOWHF_Add_c;
   		UOWHF_Add_c.7:=UOWHF_Result[7].31;
   		UOWHF_Result[7].31:=0;
   		UOWHF_Result[8]:=UOWHF_Result[8] + 1944089553+UOWHF_Add_c;
   		UOWHF_Add_c.8:=UOWHF_Result[8].31;
   		UOWHF_Result[8].31:=0;
   	End_If;
   	If UOWHF_Msg[15].[25] Then
   		UOWHF_Result[0]:=UOWHF_Result[0] + 724636145+UOWHF_Add_c;
   		UOWHF_Add_c.0:=UOWHF_Result[0].31;
   		UOWHF_Result[0].31:=0;
   		UOWHF_Result[1]:=UOWHF_Result[1] + 170859751+UOWHF_Add_c;
   		UOWHF_Add_c.1:=UOWHF_Result[1].31;
   		UOWHF_Result[1].31:=0;
   		UOWHF_Result[2]:=UOWHF_Result[2] + 155215951+UOWHF_Add_c;
   		UOWHF_Add_c.2:=UOWHF_Result[2].31;
   		UOWHF_Result[2].31:=0;
   		UOWHF_Result[3]:=UOWHF_Result[3] + 1024656956+UOWHF_Add_c;
   		UOWHF_Add_c.3:=UOWHF_Result[3].31;
   		UOWHF_Result[3].31:=0;
   		UOWHF_Result[4]:=UOWHF_Result[4] + 1793979248+UOWHF_Add_c;
   		UOWHF_Add_c.4:=UOWHF_Result[4].31;
   		UOWHF_Result[4].31:=0;
   		UOWHF_Result[5]:=UOWHF_Result[5] + 823486319+UOWHF_Add_c;
   		UOWHF_Add_c.5:=UOWHF_Result[5].31;
   		UOWHF_Result[5].31:=0;
   		UOWHF_Result[6]:=UOWHF_Result[6] + 2143852208+UOWHF_Add_c;
   		UOWHF_Add_c.6:=UOWHF_Result[6].31;
   		UOWHF_Result[6].31:=0;
   		UOWHF_Result[7]:=UOWHF_Result[7] + 2006358413+UOWHF_Add_c;
   		UOWHF_Add_c.7:=UOWHF_Result[7].31;
   		UOWHF_Result[7].31:=0;
   		UOWHF_Result[8]:=UOWHF_Result[8] + 133442244+UOWHF_Add_c;
   		UOWHF_Add_c.8:=UOWHF_Result[8].31;
   		UOWHF_Result[8].31:=0;
   	End_If;
   	If UOWHF_Msg[15].[26] Then
   		UOWHF_Result[0]:=UOWHF_Result[0] + 1586151130+UOWHF_Add_c;
   		UOWHF_Add_c.0:=UOWHF_Result[0].31;
   		UOWHF_Result[0].31:=0;
   		UOWHF_Result[1]:=UOWHF_Result[1] + 1002747430+UOWHF_Add_c;
   		UOWHF_Add_c.1:=UOWHF_Result[1].31;
   		UOWHF_Result[1].31:=0;
   		UOWHF_Result[2]:=UOWHF_Result[2] + 406974627+UOWHF_Add_c;
   		UOWHF_Add_c.2:=UOWHF_Result[2].31;
   		UOWHF_Result[2].31:=0;
   		UOWHF_Result[3]:=UOWHF_Result[3] + 1569154368+UOWHF_Add_c;
   		UOWHF_Add_c.3:=UOWHF_Result[3].31;
   		UOWHF_Result[3].31:=0;
   		UOWHF_Result[4]:=UOWHF_Result[4] + 131793540+UOWHF_Add_c;
   		UOWHF_Add_c.4:=UOWHF_Result[4].31;
   		UOWHF_Result[4].31:=0;
   		UOWHF_Result[5]:=UOWHF_Result[5] + 1162262801+UOWHF_Add_c;
   		UOWHF_Add_c.5:=UOWHF_Result[5].31;
   		UOWHF_Result[5].31:=0;
   		UOWHF_Result[6]:=UOWHF_Result[6] + 599815853+UOWHF_Add_c;
   		UOWHF_Add_c.6:=UOWHF_Result[6].31;
   		UOWHF_Result[6].31:=0;
   		UOWHF_Result[7]:=UOWHF_Result[7] + 1835326468+UOWHF_Add_c;
   		UOWHF_Add_c.7:=UOWHF_Result[7].31;
   		UOWHF_Result[7].31:=0;
   		UOWHF_Result[8]:=UOWHF_Result[8] + 1701587691+UOWHF_Add_c;
   		UOWHF_Add_c.8:=UOWHF_Result[8].31;
   		UOWHF_Result[8].31:=0;
   	End_If;
   	If UOWHF_Msg[15].[27] Then
   		UOWHF_Result[0]:=UOWHF_Result[0] + 618955582+UOWHF_Add_c;
   		UOWHF_Add_c.0:=UOWHF_Result[0].31;
   		UOWHF_Result[0].31:=0;
   		UOWHF_Result[1]:=UOWHF_Result[1] + 1664492708+UOWHF_Add_c;
   		UOWHF_Add_c.1:=UOWHF_Result[1].31;
   		UOWHF_Result[1].31:=0;
   		UOWHF_Result[2]:=UOWHF_Result[2] + 1589039931+UOWHF_Add_c;
   		UOWHF_Add_c.2:=UOWHF_Result[2].31;
   		UOWHF_Result[2].31:=0;
   		UOWHF_Result[3]:=UOWHF_Result[3] + 756852338+UOWHF_Add_c;
   		UOWHF_Add_c.3:=UOWHF_Result[3].31;
   		UOWHF_Result[3].31:=0;
   		UOWHF_Result[4]:=UOWHF_Result[4] + 1607053532+UOWHF_Add_c;
   		UOWHF_Add_c.4:=UOWHF_Result[4].31;
   		UOWHF_Result[4].31:=0;
   		UOWHF_Result[5]:=UOWHF_Result[5] + 583730900+UOWHF_Add_c;
   		UOWHF_Add_c.5:=UOWHF_Result[5].31;
   		UOWHF_Result[5].31:=0;
   		UOWHF_Result[6]:=UOWHF_Result[6] + 1552133050+UOWHF_Add_c;
   		UOWHF_Add_c.6:=UOWHF_Result[6].31;
   		UOWHF_Result[6].31:=0;
   		UOWHF_Result[7]:=UOWHF_Result[7] + 393170940+UOWHF_Add_c;
   		UOWHF_Add_c.7:=UOWHF_Result[7].31;
   		UOWHF_Result[7].31:=0;
   		UOWHF_Result[8]:=UOWHF_Result[8] + 1559800586+UOWHF_Add_c;
   		UOWHF_Add_c.8:=UOWHF_Result[8].31;
   		UOWHF_Result[8].31:=0;
   	End_If;
   	If UOWHF_Msg[15].[28] Then
   		UOWHF_Result[0]:=UOWHF_Result[0] + 1909013465+UOWHF_Add_c;
   		UOWHF_Add_c.0:=UOWHF_Result[0].31;
   		UOWHF_Result[0].31:=0;
   		UOWHF_Result[1]:=UOWHF_Result[1] + 821492496+UOWHF_Add_c;
   		UOWHF_Add_c.1:=UOWHF_Result[1].31;
   		UOWHF_Result[1].31:=0;
   		UOWHF_Result[2]:=UOWHF_Result[2] + 1496726201+UOWHF_Add_c;
   		UOWHF_Add_c.2:=UOWHF_Result[2].31;
   		UOWHF_Result[2].31:=0;
   		UOWHF_Result[3]:=UOWHF_Result[3] + 742639527+UOWHF_Add_c;
   		UOWHF_Add_c.3:=UOWHF_Result[3].31;
   		UOWHF_Result[3].31:=0;
   		UOWHF_Result[4]:=UOWHF_Result[4] + 283938920+UOWHF_Add_c;
   		UOWHF_Add_c.4:=UOWHF_Result[4].31;
   		UOWHF_Result[4].31:=0;
   		UOWHF_Result[5]:=UOWHF_Result[5] + 1599553596+UOWHF_Add_c;
   		UOWHF_Add_c.5:=UOWHF_Result[5].31;
   		UOWHF_Result[5].31:=0;
   		UOWHF_Result[6]:=UOWHF_Result[6] + 197582786+UOWHF_Add_c;
   		UOWHF_Add_c.6:=UOWHF_Result[6].31;
   		UOWHF_Result[6].31:=0;
   		UOWHF_Result[7]:=UOWHF_Result[7] + 818790931+UOWHF_Add_c;
   		UOWHF_Add_c.7:=UOWHF_Result[7].31;
   		UOWHF_Result[7].31:=0;
   		UOWHF_Result[8]:=UOWHF_Result[8] + 268526370+UOWHF_Add_c;
   		UOWHF_Add_c.8:=UOWHF_Result[8].31;
   		UOWHF_Result[8].31:=0;
   	End_If;
   	If UOWHF_Msg[15].[29] Then
   		UOWHF_Result[0]:=UOWHF_Result[0] + 1815290424+UOWHF_Add_c;
   		UOWHF_Add_c.0:=UOWHF_Result[0].31;
   		UOWHF_Result[0].31:=0;
   		UOWHF_Result[1]:=UOWHF_Result[1] + 556111681+UOWHF_Add_c;
   		UOWHF_Add_c.1:=UOWHF_Result[1].31;
   		UOWHF_Result[1].31:=0;
   		UOWHF_Result[2]:=UOWHF_Result[2] + 765690894+UOWHF_Add_c;
   		UOWHF_Add_c.2:=UOWHF_Result[2].31;
   		UOWHF_Result[2].31:=0;
   		UOWHF_Result[3]:=UOWHF_Result[3] + 200819107+UOWHF_Add_c;
   		UOWHF_Add_c.3:=UOWHF_Result[3].31;
   		UOWHF_Result[3].31:=0;
   		UOWHF_Result[4]:=UOWHF_Result[4] + 101816225+UOWHF_Add_c;
   		UOWHF_Add_c.4:=UOWHF_Result[4].31;
   		UOWHF_Result[4].31:=0;
   		UOWHF_Result[5]:=UOWHF_Result[5] + 25674087+UOWHF_Add_c;
   		UOWHF_Add_c.5:=UOWHF_Result[5].31;
   		UOWHF_Result[5].31:=0;
   		UOWHF_Result[6]:=UOWHF_Result[6] + 1692405523+UOWHF_Add_c;
   		UOWHF_Add_c.6:=UOWHF_Result[6].31;
   		UOWHF_Result[6].31:=0;
   		UOWHF_Result[7]:=UOWHF_Result[7] + 1843526161+UOWHF_Add_c;
   		UOWHF_Add_c.7:=UOWHF_Result[7].31;
   		UOWHF_Result[7].31:=0;
   		UOWHF_Result[8]:=UOWHF_Result[8] + 1561145795+UOWHF_Add_c;
   		UOWHF_Add_c.8:=UOWHF_Result[8].31;
   		UOWHF_Result[8].31:=0;
   	End_If;
   	If UOWHF_Msg[15].[30] Then
   		UOWHF_Result[0]:=UOWHF_Result[0] + 811437359+UOWHF_Add_c;
   		UOWHF_Add_c.0:=UOWHF_Result[0].31;
   		UOWHF_Result[0].31:=0;
   		UOWHF_Result[1]:=UOWHF_Result[1] + 1787609462+UOWHF_Add_c;
   		UOWHF_Add_c.1:=UOWHF_Result[1].31;
   		UOWHF_Result[1].31:=0;
   		UOWHF_Result[2]:=UOWHF_Result[2] + 823007593+UOWHF_Add_c;
   		UOWHF_Add_c.2:=UOWHF_Result[2].31;
   		UOWHF_Result[2].31:=0;
   		UOWHF_Result[3]:=UOWHF_Result[3] + 349243828+UOWHF_Add_c;
   		UOWHF_Add_c.3:=UOWHF_Result[3].31;
   		UOWHF_Result[3].31:=0;
   		UOWHF_Result[4]:=UOWHF_Result[4] + 1626029622+UOWHF_Add_c;
   		UOWHF_Add_c.4:=UOWHF_Result[4].31;
   		UOWHF_Result[4].31:=0;
   		UOWHF_Result[5]:=UOWHF_Result[5] + 1613165835+UOWHF_Add_c;
   		UOWHF_Add_c.5:=UOWHF_Result[5].31;
   		UOWHF_Result[5].31:=0;
   		UOWHF_Result[6]:=UOWHF_Result[6] + 960984991+UOWHF_Add_c;
   		UOWHF_Add_c.6:=UOWHF_Result[6].31;
   		UOWHF_Result[6].31:=0;
   		UOWHF_Result[7]:=UOWHF_Result[7] + 1552389455+UOWHF_Add_c;
   		UOWHF_Add_c.7:=UOWHF_Result[7].31;
   		UOWHF_Result[7].31:=0;
   		UOWHF_Result[8]:=UOWHF_Result[8] + 36432777+UOWHF_Add_c;
   		UOWHF_Add_c.8:=UOWHF_Result[8].31;
   		UOWHF_Result[8].31:=0;
   	End_If;
   	If UOWHF_Msg[15].[31] Then
   		UOWHF_Result[0]:=UOWHF_Result[0] + 671684221+UOWHF_Add_c;
   		UOWHF_Add_c.0:=UOWHF_Result[0].31;
   		UOWHF_Result[0].31:=0;
   		UOWHF_Result[1]:=UOWHF_Result[1] + 99804830+UOWHF_Add_c;
   		UOWHF_Add_c.1:=UOWHF_Result[1].31;
   		UOWHF_Result[1].31:=0;
   		UOWHF_Result[2]:=UOWHF_Result[2] + 1199926868+UOWHF_Add_c;
   		UOWHF_Add_c.2:=UOWHF_Result[2].31;
   		UOWHF_Result[2].31:=0;
   		UOWHF_Result[3]:=UOWHF_Result[3] + 1924295854+UOWHF_Add_c;
   		UOWHF_Add_c.3:=UOWHF_Result[3].31;
   		UOWHF_Result[3].31:=0;
   		UOWHF_Result[4]:=UOWHF_Result[4] + 196799211+UOWHF_Add_c;
   		UOWHF_Add_c.4:=UOWHF_Result[4].31;
   		UOWHF_Result[4].31:=0;
   		UOWHF_Result[5]:=UOWHF_Result[5] + 892312821+UOWHF_Add_c;
   		UOWHF_Add_c.5:=UOWHF_Result[5].31;
   		UOWHF_Result[5].31:=0;
   		UOWHF_Result[6]:=UOWHF_Result[6] + 1548504499+UOWHF_Add_c;
   		UOWHF_Add_c.6:=UOWHF_Result[6].31;
   		UOWHF_Result[6].31:=0;
   		UOWHF_Result[7]:=UOWHF_Result[7] + 1330003781+UOWHF_Add_c;
   		UOWHF_Add_c.7:=UOWHF_Result[7].31;
   		UOWHF_Result[7].31:=0;
   		UOWHF_Result[8]:=UOWHF_Result[8] + 1711999757+UOWHF_Add_c;
   		UOWHF_Add_c.8:=UOWHF_Result[8].31;
   		UOWHF_Result[8].31:=0;
   	End_If;
   		UOWHF_Result[UOWHF_OutputMaxInd]:=UOWHF_Result[UOWHF_OutputMaxInd] and 16#FFF; //clear high bit
   *)
END_ROUTINE

ROUTINE UOWHF_Init   (* structured text *)
   Case UOWHF_Ver OF
   0:
   	UOWHF_InputLen:=255;  //bits of input.
   	UOWHF_InputMaxInd:=8;  //maximum index for dints which store the bits of input.
    	For UOWHF_i:=0 to UOWHF_InputMaxInd by 1 do
   		UOWHF_Result[UOWHF_i]:=0;
   	End_For;
   1:
   	UOWHF_InputLen:= 383;
   	UOWHF_InputMaxInd:=12;  //maximum index for array.
    	For UOWHF_i:=0 to UOWHF_InputMaxInd by 1 do
   		UOWHF_Result[UOWHF_i]:=0;
   	End_For;
   2:
   	UOWHF_InputLen:= 511;
   	UOWHF_InputMaxInd:=16;  //maximum index for array.
   	 For UOWHF_i:=0 to UOWHF_InputMaxInd by 1 do
   		UOWHF_Result[UOWHF_i]:=0;
   	End_For;
   End_Case;
   
   UOWHF_OutputMaxInd := UOWHF_InputMaxInd/2;
END_ROUTINE

ROUTINE UOWHF_Test   (* structured text *)
   //Description: initialize the variables.
   
   
   UOWHF_Ver:=2;
   
   UOWHF_Vary_MsgLen:=17;
   
   if S:FS then  (* this is the first, normal scan of the routines in the current program, initialize the program.*)
   	 //UOWHF_Ver means that the version of OWF: 256-256 bits, 384-384 bits, and 512-512 bits. The first number is length of input, the last number is length of output.
                    //If UOWHF_Ver means that the version of Hash, then three versions are: 256-128 bits, 384-160 bits and 512-256 bits.
   	If UOWHF_Ver=0 then
   		for UOWHF_i:=0 to UOWHF_Vary_MsgLen by 1 Do
   			UOWHF_Vary_Message[UOWHF_i]:= 65535;   //Half of the selection factors are 1.
   			//UOWHF_Msg[UOWHF_i]:= -1;    //All the selection factors are 1.
   		end_for;
   	end_if;
   
   	If UOWHF_Ver=1 then
   		for UOWHF_i:=0 to UOWHF_Vary_MsgLen by 1 Do
   			UOWHF_Vary_Message[UOWHF_i]:= 65535;     //Half of the selection factors are 1.
   			//UOWHF_Msg[UOWHF_i]:= -1;   //All the selection factors are 1.
   		end_for;
   	end_if;
   
   	If UOWHF_Ver=2 then
   		for UOWHF_i:=0 to UOWHF_Vary_MsgLen by 1 Do
   			UOWHF_Vary_Message[UOWHF_i]:= 65535;     //Half of the selection factors are 1.
   			//UOWHF_Msg[UOWHF_i]:= -1;   //All the selection factors are 1.
   		end_for;
   	end_if;
   
   end_if;
   
   jsr(UOWHF_Vary);
   
   
   
   
END_ROUTINE

ROUTINE UOWHF_Vary   (* structured text *)
   
   
   JSR(UOWHF_Init);
   
   
   UOWHF_VaryLen:=(UOWHF_Vary_MsgLen+1) MOD (UOWHF_OutputMaxInd+1);
   If UOWHF_VaryLen<>0 Then
   	UOWHF_VaryLen:=UOWHF_OutputMaxInd+1 - UOWHF_VaryLen;
   
   	//pad 1 if neccessary
   	For UOWHF_Vary_i:=UOWHF_Vary_MsgLen+1 to UOWHF_Vary_MsgLen+UOWHF_VaryLen by 1 Do
   
   		UOWHF_Vary_Message[UOWHF_Vary_i]:=65535;
   
   	End_For;
   	UOWHF_Vary_MsgLen:=UOWHF_Vary_MsgLen+UOWHF_VaryLen;
   End_if;
   
   
   UOWHF_Vary_BlkNum:= (UOWHF_Vary_MsgLen+1)/(UOWHF_OutputMaxInd+1)-1 ;
   
   For UOWHF_Vary_i:=0 to UOWHF_InputMaxInd by 1 Do
   	UOWHF_Msg[UOWHF_Vary_i]:=UOWHF_Vary_Message[UOWHF_Vary_i];
   End_For;
   JSR(UOWHF);
   
   UOWHF_Vary_z:=UOWHF_InputMaxInd+1;
   For UOWHF_Vary_i:=2 to UOWHF_Vary_BlkNum by 1 Do
   
   	For UOWHF_Vary_j:=0 to UOWHF_OutputMaxInd by 1 Do
   		UOWHF_Msg[UOWHF_Vary_j]:=UOWHF_Vary_Message[UOWHF_Vary_z+UOWHF_Vary_j];
   		UOWHF_Msg[UOWHF_Vary_j+UOWHF_OutputMaxInd+1]:=UOWHF_Result[UOWHF_Vary_j];
   	End_For;
   	JSR(UOWHF);
   	UOWHF_Vary_z:=UOWHF_Vary_z+UOWHF_OutputMaxInd+1;
   End_For;
   
   
   
END_ROUTINE
END_PROGRAM
